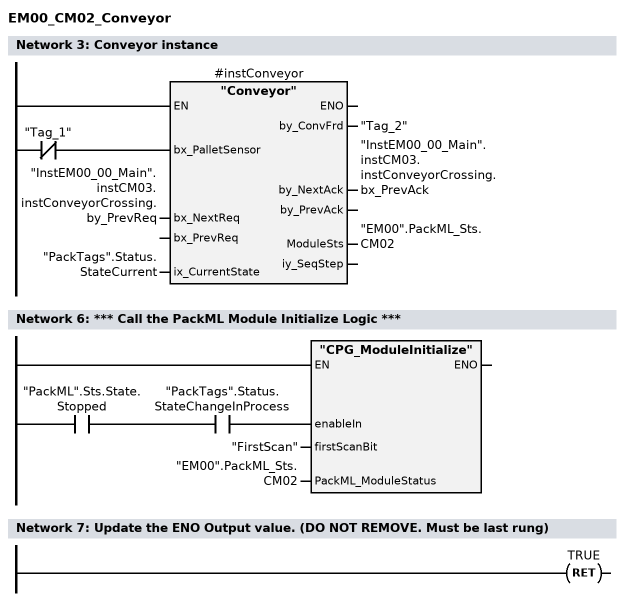
   RUNG wire#powerrail
      #instConveyor(bx_PalletSensor := wire#w1, bx_NextReq := "InstEM00_00_Main".instCM03.instConveyorCrossing.by_PrevReq, bx_PrevReq :=, ix_CurrentState := "PackTags".Status.StateCurrent, by_ConvFrd => "Tag_2", by_NextAck => "InstEM00_00_Main".instCM03.instConveyorCrossing.bx_PrevAck, by_PrevAck =>, ModuleSts => "EM00".PackML_Sts.CM02, iy_SeqStep =>)
   END_RUNG
   RUNG wire#powerrail
      I_Contact( "Tag_1" )
   END_RUNG wire#w1
   // the same network as SCL:
   #instConveyor(bx_PalletSensor := NOT "Tag_1",   // "Conveyor"
                 bx_NextReq := "InstEM00_00_Main".instCM03.instConveyorCrossing.by_PrevReq,
                 ix_CurrentState := "PackTags".Status.StateCurrent,
                 by_ConvFrd => "Tag_2",
                 by_NextAck => "InstEM00_00_Main".instCM03.instConveyorCrossing.bx_PrevAck,
                 ModuleSts => "EM00".PackML_Sts.CM02);
END_REGION

REGION Network 4: *** Begin the Event Information Section ***
END_REGION

REGION Network 5: *** Begin the State Model Status Feedback Section ***
END_REGION

REGION Network 6: *** Call the PackML Module Initialize Logic ***
   RUNG wire#powerrail
      "CPG_ModuleInitialize"(enableIn := wire#w1, firstScanBit := "FirstScan", PackML_ModuleStatus := "EM00".PackML_Sts.CM02)
   END_RUNG
   RUNG wire#powerrail
      Contact( "PackML".Sts.State.Stopped )
      Contact( "PackTags".Status.StateChangeInProcess )
   END_RUNG wire#w1
   // the same network as SCL:
   "CPG_ModuleInitialize"(enableIn := "PackML".Sts.State.Stopped AND "PackTags".Status.StateChangeInProcess,
                          firstScanBit := "FirstScan",
                          PackML_ModuleStatus := "EM00".PackML_Sts.CM02);
END_REGION

REGION Network 7: Update the ENO Output value. (DO NOT REMOVE. Must be last rung)
   RUNG wire#powerrail
      ReturnCoil( TRUE )
   END_RUNG
   // the same network as SCL:
   ENO := TRUE;
   RETURN;
END_REGION
END_FUNCTION_BLOCK

FUNCTION_BLOCK "EM00_CM03_ConveyorCrossing"   // FB31653, LAD
TITLE = EM00_CM03
{ S7_Optimized_Access := 'TRUE' }
AUTHOR : tech.team.motioncontrol@siemens.com
FAMILY : CPG
VERSION : 1.1
// Support: tech.team.motioncontrol@siemens.com
   VAR
      statDummyBool : Bool;   // dummy bool - placeholder
      instConveyorCrossing : "ConveyorCrossing";
   END_VAR
BEGIN

REGION Network 1: *** Begin the Setpoint Management Information Section ***
END_REGION

REGION Network 2: *** Begin the Logic Section ***
END_REGION

REGION Network 3: Conveyor crossing instance
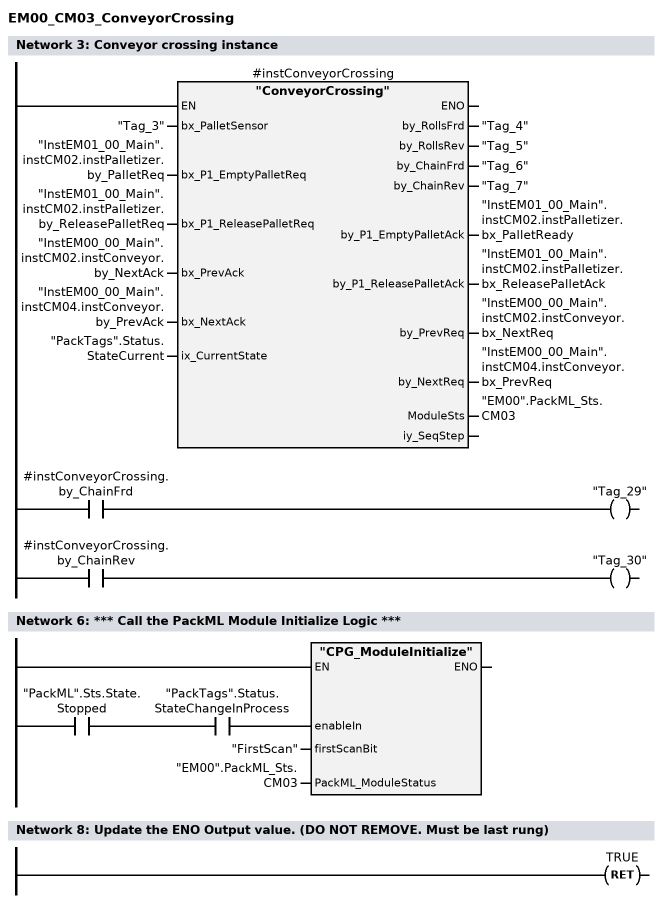
   RUNG wire#powerrail
      #instConveyorCrossing(bx_PalletSensor := "Tag_3", bx_P1_EmptyPalletReq := "InstEM01_00_Main".instCM02.instPalletizer.by_PalletReq, bx_P1_ReleasePalletReq := "InstEM01_00_Main".instCM02.instPalletizer.by_ReleasePalletReq, bx_PrevAck := "InstEM00_00_Main".instCM02.instConveyor.by_NextAck, bx_NextAck := "InstEM00_00_Main".instCM04.instConveyor.by_PrevAck, ix_CurrentState := "PackTags".Status.StateCurrent, by_RollsFrd => "Tag_4", by_RollsRev => "Tag_5", by_ChainFrd => "Tag_6", by_ChainRev => "Tag_7", by_P1_EmptyPalletAck => "InstEM01_00_Main".instCM02.instPalletizer.bx_PalletReady, by_P1_ReleasePalletAck => "InstEM01_00_Main".instCM02.instPalletizer.bx_ReleasePalletAck, by_PrevReq => "InstEM00_00_Main".instCM02.instConveyor.bx_NextReq, by_NextReq => "InstEM00_00_Main".instCM04.instConveyor.bx_PrevReq, ModuleSts => "EM00".PackML_Sts.CM03, iy_SeqStep =>)
   END_RUNG
   RUNG wire#powerrail
      Contact( #instConveyorCrossing.by_ChainFrd )
      Coil( "Tag_29" )
   END_RUNG
   RUNG wire#powerrail
      Contact( #instConveyorCrossing.by_ChainRev )
      Coil( "Tag_30" )
   END_RUNG
   // the same network as SCL:
   #instConveyorCrossing(bx_PalletSensor := "Tag_3",   // "ConveyorCrossing"
                         bx_P1_EmptyPalletReq := "InstEM01_00_Main".instCM02.instPalletizer.by_PalletReq,
                         bx_P1_ReleasePalletReq := "InstEM01_00_Main".instCM02.instPalletizer.by_ReleasePalletReq,
                         bx_PrevAck := "InstEM00_00_Main".instCM02.instConveyor.by_NextAck,
                         bx_NextAck := "InstEM00_00_Main".instCM04.instConveyor.by_PrevAck,
                         ix_CurrentState := "PackTags".Status.StateCurrent,
                         by_RollsFrd => "Tag_4",
                         by_RollsRev => "Tag_5",
                         by_ChainFrd => "Tag_6",
                         by_ChainRev => "Tag_7",
                         by_P1_EmptyPalletAck => "InstEM01_00_Main".instCM02.instPalletizer.bx_PalletReady,
                         by_P1_ReleasePalletAck => "InstEM01_00_Main".instCM02.instPalletizer.bx_ReleasePalletAck,
                         by_PrevReq => "InstEM00_00_Main".instCM02.instConveyor.bx_NextReq,
                         by_NextReq => "InstEM00_00_Main".instCM04.instConveyor.bx_PrevReq,
                         ModuleSts => "EM00".PackML_Sts.CM03);
   "Tag_29" := #instConveyorCrossing.by_ChainFrd;
   "Tag_30" := #instConveyorCrossing.by_ChainRev;
END_REGION

REGION Network 4: *** Begin the Event Information Section ***
END_REGION

REGION Network 5: *** Begin the State Model Status Feedback Section ***
END_REGION

REGION Network 6: *** Call the PackML Module Initialize Logic ***
   RUNG wire#powerrail
      "CPG_ModuleInitialize"(enableIn := wire#w1, firstScanBit := "FirstScan", PackML_ModuleStatus := "EM00".PackML_Sts.CM03)
   END_RUNG
   RUNG wire#powerrail
      Contact( "PackML".Sts.State.Stopped )
      Contact( "PackTags".Status.StateChangeInProcess )
   END_RUNG wire#w1
   // the same network as SCL:
   "CPG_ModuleInitialize"(enableIn := "PackML".Sts.State.Stopped AND "PackTags".Status.StateChangeInProcess,
                          firstScanBit := "FirstScan",
                          PackML_ModuleStatus := "EM00".PackML_Sts.CM03);
END_REGION

REGION Network 8: Update the ENO Output value. (DO NOT REMOVE. Must be last rung)
   RUNG wire#powerrail
      ReturnCoil( TRUE )
   END_RUNG
   // the same network as SCL:
   ENO := TRUE;
   RETURN;
END_REGION
END_FUNCTION_BLOCK

FUNCTION_BLOCK "EM00_CM04_Conveyor"   // FB31654, LAD
TITLE = EM00_CM04
{ S7_Optimized_Access := 'TRUE' }
AUTHOR : tech.team.motioncontrol@siemens.com
FAMILY : CPG
VERSION : 1.1
// Support: tech.team.motioncontrol@siemens.com
   VAR
      statDummyBool : Bool;   // dummy bool - placeholder
      instConveyor : "Conveyor";
   END_VAR
BEGIN

REGION Network 1: *** Begin the Setpoint Management Information Section ***
END_REGION

REGION Network 2: *** Begin the Logic Section ***
END_REGION

REGION Network 3: Conveyor instance
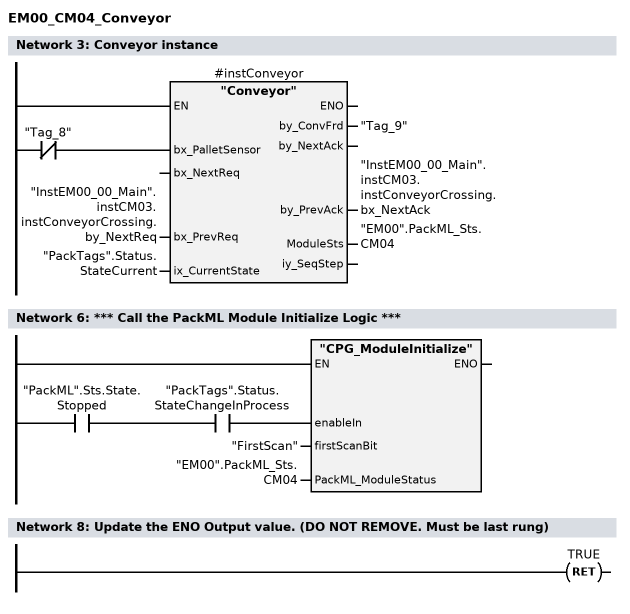
   RUNG wire#powerrail
      #instConveyor(bx_PalletSensor := wire#w1, bx_NextReq :=, bx_PrevReq := "InstEM00_00_Main".instCM03.instConveyorCrossing.by_NextReq, ix_CurrentState := "PackTags".Status.StateCurrent, by_ConvFrd => "Tag_9", by_NextAck =>, by_PrevAck => "InstEM00_00_Main".instCM03.instConveyorCrossing.bx_NextAck, ModuleSts => "EM00".PackML_Sts.CM04, iy_SeqStep =>)
   END_RUNG
   RUNG wire#powerrail
      I_Contact( "Tag_8" )
   END_RUNG wire#w1
   // the same network as SCL:
   #instConveyor(bx_PalletSensor := NOT "Tag_8",   // "Conveyor"
                 bx_PrevReq := "InstEM00_00_Main".instCM03.instConveyorCrossing.by_NextReq,
                 ix_CurrentState := "PackTags".Status.StateCurrent,
                 by_ConvFrd => "Tag_9",
                 by_PrevAck => "InstEM00_00_Main".instCM03.instConveyorCrossing.bx_NextAck,
                 ModuleSts => "EM00".PackML_Sts.CM04);
END_REGION

REGION Network 4: *** Begin the Event Information Section ***
END_REGION

REGION Network 5: *** Begin the State Model Status Feedback Section ***
END_REGION

REGION Network 6: *** Call the PackML Module Initialize Logic ***
   RUNG wire#powerrail
      "CPG_ModuleInitialize"(enableIn := wire#w1, firstScanBit := "FirstScan", PackML_ModuleStatus := "EM00".PackML_Sts.CM04)
   END_RUNG
   RUNG wire#powerrail
      Contact( "PackML".Sts.State.Stopped )
      Contact( "PackTags".Status.StateChangeInProcess )
   END_RUNG wire#w1
   // the same network as SCL:
   "CPG_ModuleInitialize"(enableIn := "PackML".Sts.State.Stopped AND "PackTags".Status.StateChangeInProcess,
                          firstScanBit := "FirstScan",
                          PackML_ModuleStatus := "EM00".PackML_Sts.CM04);
END_REGION

REGION Network 8: Update the ENO Output value. (DO NOT REMOVE. Must be last rung)
   RUNG wire#powerrail
      ReturnCoil( TRUE )
   END_RUNG
   // the same network as SCL:
   ENO := TRUE;
   RETURN;
END_REGION
END_FUNCTION_BLOCK

FUNCTION_BLOCK "EM00_CM05_ConveyorCrossing"   // FB31655, LAD
TITLE = EM00_CM05
{ S7_Optimized_Access := 'TRUE' }
AUTHOR : tech.team.motioncontrol@siemens.com
FAMILY : CPG
VERSION : 1.1
// Support: tech.team.motioncontrol@siemens.com
   VAR
      statDummyBool : Bool;   // dummy bool - placeholder
   END_VAR
BEGIN

REGION Network 1: *** Begin the Setpoint Management Information Section ***
END_REGION

REGION Network 2: *** Begin the Logic Section ***
END_REGION

REGION Network 3: *** Begin the Event Information Section ***
END_REGION

REGION Network 4: *** Begin the State Model Status Feedback Section ***
END_REGION

REGION Network 5: *** Call the PackML Module Initialize Logic ***
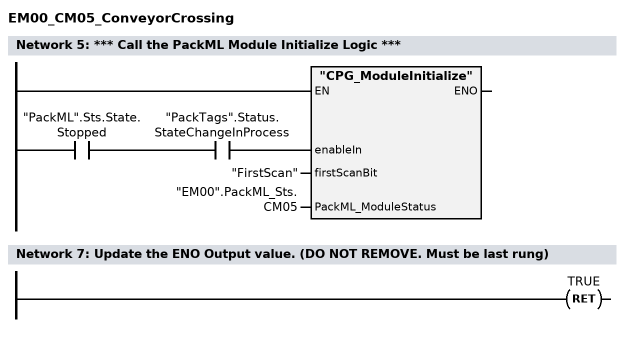
   RUNG wire#powerrail
      "CPG_ModuleInitialize"(enableIn := wire#w1, firstScanBit := "FirstScan", PackML_ModuleStatus := "EM00".PackML_Sts.CM05)
   END_RUNG
   RUNG wire#powerrail
      Contact( "PackML".Sts.State.Stopped )
      Contact( "PackTags".Status.StateChangeInProcess )
   END_RUNG wire#w1
   // the same network as SCL:
   "CPG_ModuleInitialize"(enableIn := "PackML".Sts.State.Stopped AND "PackTags".Status.StateChangeInProcess,
                          firstScanBit := "FirstScan",
                          PackML_ModuleStatus := "EM00".PackML_Sts.CM05);
END_REGION

REGION Network 7: Update the ENO Output value. (DO NOT REMOVE. Must be last rung)
   RUNG wire#powerrail
      ReturnCoil( TRUE )
   END_RUNG
   // the same network as SCL:
   ENO := TRUE;
   RETURN;
END_REGION
END_FUNCTION_BLOCK

// folder: EM01_Palletizing

FUNCTION_BLOCK "EM01_00_Main"   // FB31660, LAD
TITLE = EM01_00_Main
{ S7_Optimized_Access := 'TRUE' }
AUTHOR : tech.team.motioncontrol@siemens.com
FAMILY : CPG
VERSION : 1.1
// Support: tech.team.motioncontrol@siemens.com
   VAR
      instEventControl : "EM01_01_EventControl";   // Instance DB - EM's Event Control Logic
      instPackML_ModuleSum : "EM01_02_PackML_ModuleSum";   // Instance DB - EM's PackML Module Summation Logic
      instCM01 : "EM01_CM01_Conveyor";   // Instance DB - CM01
      instCM02 : "EM01_CM02_Palletizer";   // Instance DB - CM02
   END_VAR
   VAR_TEMP   // added for the SCL form of the ladder/FBD networks
      _w1 : Bool;
   END_VAR
BEGIN

REGION Network 1: *** BEGIN MAIN LOGIC SECTION ***
END_REGION

REGION Network 2: Call the Control Module Logic - CM01
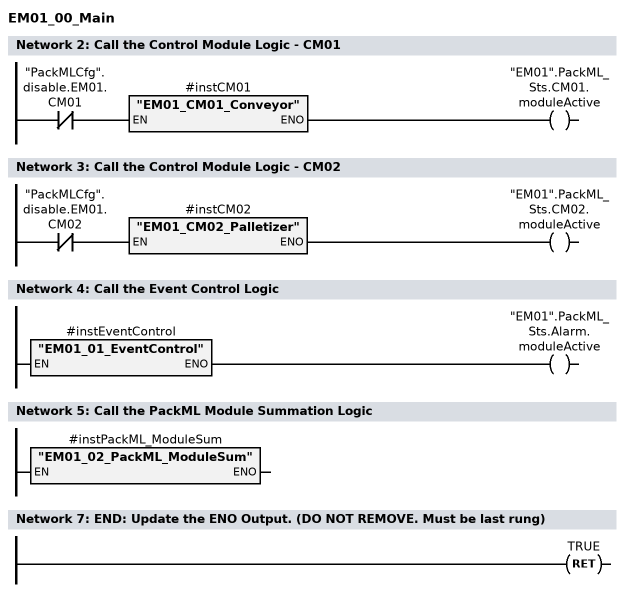
   RUNG wire#powerrail
      I_Contact( "PackMLCfg".disable.EM01.CM01 )
      #instCM01()
      Coil( "EM01".PackML_Sts.CM01.moduleActive )
   END_RUNG
   // the same network as SCL:
   #instCM01(EN := NOT "PackMLCfg".disable.EM01.CM01, ENO => #_w1);   // "EM01_CM01_Conveyor"
   "EM01".PackML_Sts.CM01.moduleActive := #_w1;
END_REGION

REGION Network 3: Call the Control Module Logic - CM02
   RUNG wire#powerrail
      I_Contact( "PackMLCfg".disable.EM01.CM02 )
      #instCM02()
      Coil( "EM01".PackML_Sts.CM02.moduleActive )
   END_RUNG
   // the same network as SCL:
   #instCM02(EN := NOT "PackMLCfg".disable.EM01.CM02, ENO => #_w1);   // "EM01_CM02_Palletizer"
   "EM01".PackML_Sts.CM02.moduleActive := #_w1;
END_REGION

REGION Network 4: Call the Event Control Logic
   RUNG wire#powerrail
      #instEventControl()
      Coil( "EM01".PackML_Sts.Alarm.moduleActive )
   END_RUNG
   // the same network as SCL:
   #instEventControl(ENO => #_w1);   // "EM01_01_EventControl"
   "EM01".PackML_Sts.Alarm.moduleActive := #_w1;
END_REGION

REGION Network 5: Call the PackML Module Summation Logic
   RUNG wire#powerrail
      #instPackML_ModuleSum()
   END_RUNG
   // the same network as SCL:
   #instPackML_ModuleSum();   // "EM01_02_PackML_ModuleSum"
END_REGION

REGION Network 7: END: Update the ENO Output. (DO NOT REMOVE. Must be last rung)
   RUNG wire#powerrail
      ReturnCoil( TRUE )
   END_RUNG
   // the same network as SCL:
   ENO := TRUE;
   RETURN;
END_REGION
END_FUNCTION_BLOCK

FUNCTION_BLOCK "EM01_01_EventControl"   // FB31661, LAD
TITLE = EM01_01_EventControl
{ S7_Optimized_Access := 'TRUE' }
AUTHOR : tech.team.motioncontrol@siemens.com
FAMILY : CPG
VERSION : 1.1
// Support: tech.team.motioncontrol@siemens.com
   VAR
      instEventMgr_Alarm : "CPG_EventManager";   // instance FB - Event Manager - Alarm Events
      instEventMgr_Warning : "CPG_EventManager";   // instance FB - Event Manager - Warning Events
      instEventMgr_Status : "CPG_EventManager";   // instance FB - Event Manager - Status Events
      instStatus_AlarmNotReset : "CPG_Event";   // instance FB - PackML Event - Alarms not reset
      statEventMgr_Cmd_Reset : Bool;   // Reset Cmd for all event managers
      statEventMgr_Cmd_Clear1stFlt : Bool;   // Clear 1st Fault Cmd for all event managers
      statEventMgr_Clear1stFlt_OS : Bool;   // Clear 1st Fault Cmd - One shot
   END_VAR
   VAR_TEMP   // added for the SCL form of the ladder/FBD networks
      _w1 : Bool;
      _w2 : Bool;
   END_VAR
BEGIN

REGION Network 1: ** STATE MODEL REPORTING STATUS ****
END_REGION

REGION Network 2: *** Call the PackML Module Initialize Logic ***
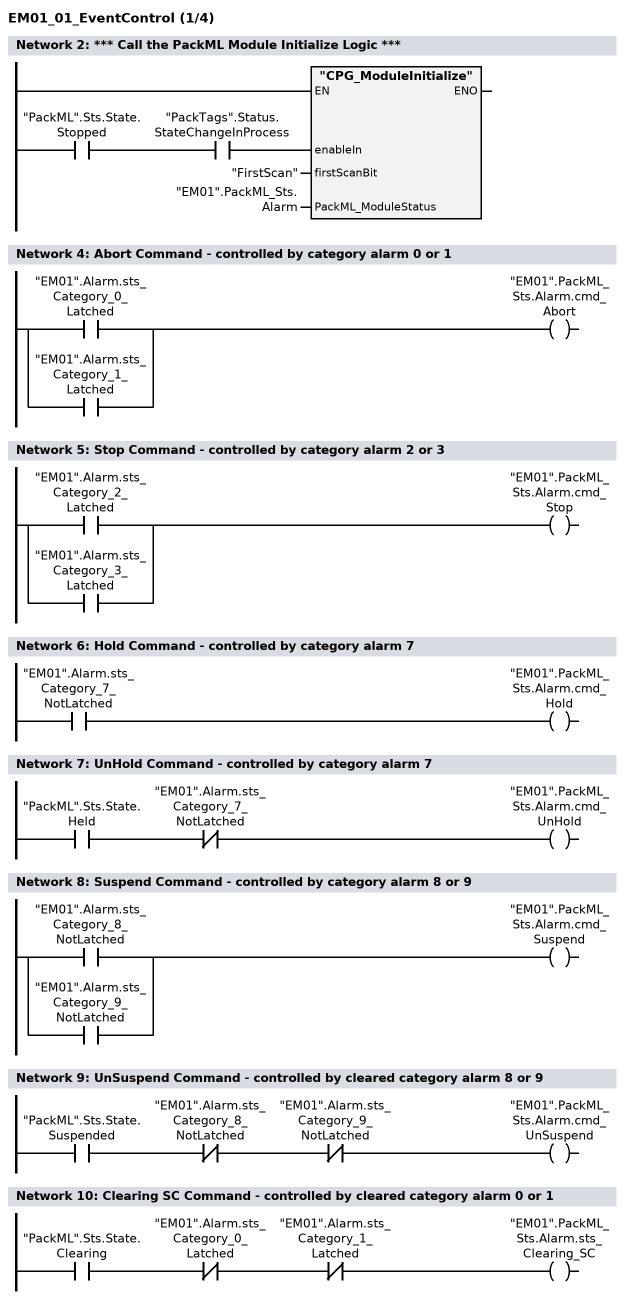
   RUNG wire#powerrail
      "CPG_ModuleInitialize"(enableIn := wire#w1, firstScanBit := "FirstScan", PackML_ModuleStatus := "EM01".PackML_Sts.Alarm)
   END_RUNG
   RUNG wire#powerrail
      Contact( "PackML".Sts.State.Stopped )
      Contact( "PackTags".Status.StateChangeInProcess )
   END_RUNG wire#w1
   // the same network as SCL:
   "CPG_ModuleInitialize"(enableIn := "PackML".Sts.State.Stopped AND "PackTags".Status.StateChangeInProcess,
                          firstScanBit := "FirstScan",
                          PackML_ModuleStatus := "EM01".PackML_Sts.Alarm);
END_REGION

REGION Network 3: Begin the LOGIC section.
END_REGION

REGION Network 4: Abort Command - controlled by category alarm 0 or 1
   RUNG wire#powerrail
      Contact( "EM01".Alarm.sts_Category_0_Latched )
      wire#w1
      Coil( "EM01".PackML_Sts.Alarm.cmd_Abort )
   END_RUNG
   RUNG wire#powerrail
      Contact( "EM01".Alarm.sts_Category_1_Latched )
   END_RUNG wire#w1
   // the same network as SCL:
   "EM01".PackML_Sts.Alarm.cmd_Abort := "EM01".Alarm.sts_Category_0_Latched OR "EM01".Alarm.sts_Category_1_Latched;
END_REGION

REGION Network 5: Stop Command - controlled by category alarm 2 or 3
   RUNG wire#powerrail
      Contact( "EM01".Alarm.sts_Category_2_Latched )
      wire#w1
      Coil( "EM01".PackML_Sts.Alarm.cmd_Stop )
   END_RUNG
   RUNG wire#powerrail
      Contact( "EM01".Alarm.sts_Category_3_Latched )
   END_RUNG wire#w1
   // the same network as SCL:
   "EM01".PackML_Sts.Alarm.cmd_Stop := "EM01".Alarm.sts_Category_2_Latched OR "EM01".Alarm.sts_Category_3_Latched;
END_REGION

REGION Network 6: Hold Command - controlled by category alarm 7
   RUNG wire#powerrail
      Contact( "EM01".Alarm.sts_Category_7_NotLatched )
      Coil( "EM01".PackML_Sts.Alarm.cmd_Hold )
   END_RUNG
   // the same network as SCL:
   "EM01".PackML_Sts.Alarm.cmd_Hold := "EM01".Alarm.sts_Category_7_NotLatched;
END_REGION

REGION Network 7: UnHold Command - controlled by category alarm 7
   RUNG wire#powerrail
      Contact( "PackML".Sts.State.Held )
      I_Contact( "EM01".Alarm.sts_Category_7_NotLatched )
      Coil( "EM01".PackML_Sts.Alarm.cmd_UnHold )
   END_RUNG
   // the same network as SCL:
   "EM01".PackML_Sts.Alarm.cmd_UnHold := "PackML".Sts.State.Held AND NOT "EM01".Alarm.sts_Category_7_NotLatched;
END_REGION

REGION Network 8: Suspend Command - controlled by category alarm 8 or 9
   RUNG wire#powerrail
      Contact( "EM01".Alarm.sts_Category_8_NotLatched )
      wire#w1
      Coil( "EM01".PackML_Sts.Alarm.cmd_Suspend )
   END_RUNG
   RUNG wire#powerrail
      Contact( "EM01".Alarm.sts_Category_9_NotLatched )
   END_RUNG wire#w1
   // the same network as SCL:
   "EM01".PackML_Sts.Alarm.cmd_Suspend := "EM01".Alarm.sts_Category_8_NotLatched OR "EM01".Alarm.sts_Category_9_NotLatched;
END_REGION

REGION Network 9: UnSuspend Command - controlled by cleared category alarm 8 or 9
   RUNG wire#powerrail
      Contact( "PackML".Sts.State.Suspended )
      I_Contact( "EM01".Alarm.sts_Category_8_NotLatched )
      I_Contact( "EM01".Alarm.sts_Category_9_NotLatched )
      Coil( "EM01".PackML_Sts.Alarm.cmd_UnSuspend )
   END_RUNG
   // the same network as SCL:
   "EM01".PackML_Sts.Alarm.cmd_UnSuspend := "PackML".Sts.State.Suspended AND NOT "EM01".Alarm.sts_Category_8_NotLatched AND NOT "EM01".Alarm.sts_Category_9_NotLatched;
END_REGION

REGION Network 10: Clearing SC Command - controlled by cleared category alarm 0 or 1
   RUNG wire#powerrail
      Contact( "PackML".Sts.State.Clearing )
      I_Contact( "EM01".Alarm.sts_Category_0_Latched )
      I_Contact( "EM01".Alarm.sts_Category_1_Latched )
      Coil( "EM01".PackML_Sts.Alarm.sts_Clearing_SC )
   END_RUNG
   // the same network as SCL:
   "EM01".PackML_Sts.Alarm.sts_Clearing_SC := "PackML".Sts.State.Clearing AND NOT "EM01".Alarm.sts_Category_0_Latched AND NOT "EM01".Alarm.sts_Category_1_Latched;
END_REGION

REGION Network 11: Resetting SC Command - controlled by cleared category alarm 0-3
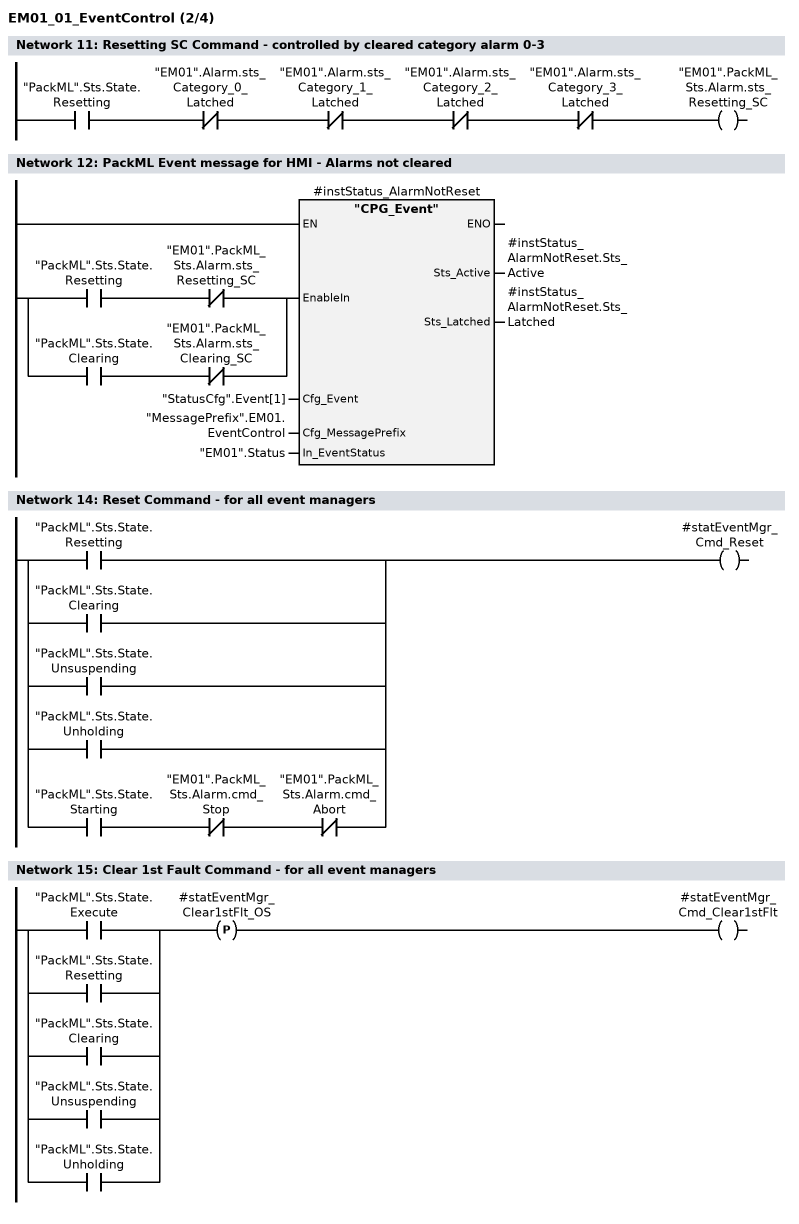
   RUNG wire#powerrail
      Contact( "PackML".Sts.State.Resetting )
      I_Contact( "EM01".Alarm.sts_Category_0_Latched )
      I_Contact( "EM01".Alarm.sts_Category_1_Latched )
      I_Contact( "EM01".Alarm.sts_Category_2_Latched )
      I_Contact( "EM01".Alarm.sts_Category_3_Latched )
      Coil( "EM01".PackML_Sts.Alarm.sts_Resetting_SC )
   END_RUNG
   // the same network as SCL:
   "EM01".PackML_Sts.Alarm.sts_Resetting_SC := "PackML".Sts.State.Resetting AND NOT "EM01".Alarm.sts_Category_0_Latched AND NOT "EM01".Alarm.sts_Category_1_Latched AND NOT "EM01".Alarm.sts_Category_2_Latched AND NOT "EM01".Alarm.sts_Category_3_Latched;
END_REGION

REGION Network 12: PackML Event message for HMI - Alarms not cleared
   RUNG wire#powerrail
      #instStatus_AlarmNotReset(EnableIn := wire#w1, Cfg_Event := "StatusCfg".Event[1], Cfg_MessagePrefix := "MessagePrefix".EM01.EventControl, In_EventStatus := "EM01".Status, Sts_Active => #instStatus_AlarmNotReset.Sts_Active, Sts_Latched => #instStatus_AlarmNotReset.Sts_Latched)
   END_RUNG
   RUNG wire#powerrail
      Contact( "PackML".Sts.State.Resetting )
      I_Contact( "EM01".PackML_Sts.Alarm.sts_Resetting_SC )
   END_RUNG wire#w1
   RUNG wire#powerrail
      Contact( "PackML".Sts.State.Clearing )
      I_Contact( "EM01".PackML_Sts.Alarm.sts_Clearing_SC )
   END_RUNG wire#w1
   // the same network as SCL:
   #instStatus_AlarmNotReset(EnableIn := ("PackML".Sts.State.Resetting AND NOT "EM01".PackML_Sts.Alarm.sts_Resetting_SC) OR ("PackML".Sts.State.Clearing AND NOT "EM01".PackML_Sts.Alarm.sts_Clearing_SC),   // "CPG_Event"
                           Cfg_Event := "StatusCfg".Event[1],
                           Cfg_MessagePrefix := "MessagePrefix".EM01.EventControl,
                           In_EventStatus := "EM01".Status,
                           Sts_Active => #instStatus_AlarmNotReset.Sts_Active,
                           Sts_Latched => #instStatus_AlarmNotReset.Sts_Latched);
END_REGION

REGION Network 13: *** EVENT CONTROL MANAGERS ***
END_REGION

REGION Network 14: Reset Command - for all event managers
   RUNG wire#powerrail
      Contact( "PackML".Sts.State.Resetting )
      wire#w1
      Coil( #statEventMgr_Cmd_Reset )
   END_RUNG
   RUNG wire#powerrail
      Contact( "PackML".Sts.State.Clearing )
   END_RUNG wire#w1
   RUNG wire#powerrail
      Contact( "PackML".Sts.State.Unsuspending )
   END_RUNG wire#w1
   RUNG wire#powerrail
      Contact( "PackML".Sts.State.Unholding )
   END_RUNG wire#w1
   RUNG wire#powerrail
      Contact( "PackML".Sts.State.Starting )
      I_Contact( "EM01".PackML_Sts.Alarm.cmd_Stop )
      I_Contact( "EM01".PackML_Sts.Alarm.cmd_Abort )
   END_RUNG wire#w1
   // the same network as SCL:
   #statEventMgr_Cmd_Reset := "PackML".Sts.State.Resetting OR "PackML".Sts.State.Clearing OR "PackML".Sts.State.Unsuspending OR "PackML".Sts.State.Unholding OR ("PackML".Sts.State.Starting AND NOT "EM01".PackML_Sts.Alarm.cmd_Stop AND NOT "EM01".PackML_Sts.Alarm.cmd_Abort);
END_REGION

REGION Network 15: Clear 1st Fault Command - for all event managers
   RUNG wire#powerrail
      Contact( "PackML".Sts.State.Execute )
      wire#w1
      P_Trig( #statEventMgr_Clear1stFlt_OS )
      Coil( #statEventMgr_Cmd_Clear1stFlt )
   END_RUNG
   RUNG wire#powerrail
      Contact( "PackML".Sts.State.Resetting )
   END_RUNG wire#w1
   RUNG wire#powerrail
      Contact( "PackML".Sts.State.Clearing )
   END_RUNG wire#w1
   RUNG wire#powerrail
      Contact( "PackML".Sts.State.Unsuspending )
   END_RUNG wire#w1
   RUNG wire#powerrail
      Contact( "PackML".Sts.State.Unholding )
   END_RUNG wire#w1
   // the same network as SCL:
   #_w1 := "PackML".Sts.State.Execute OR "PackML".Sts.State.Resetting OR "PackML".Sts.State.Clearing OR "PackML".Sts.State.Unsuspending OR "PackML".Sts.State.Unholding;
   #_w2 := #_w1 AND NOT #statEventMgr_Clear1stFlt_OS;   // rising edge
   #statEventMgr_Clear1stFlt_OS := #_w1;
   #statEventMgr_Cmd_Clear1stFlt := #_w2;
END_REGION

REGION Network 16: Call the Event Manager logic for EM alarms
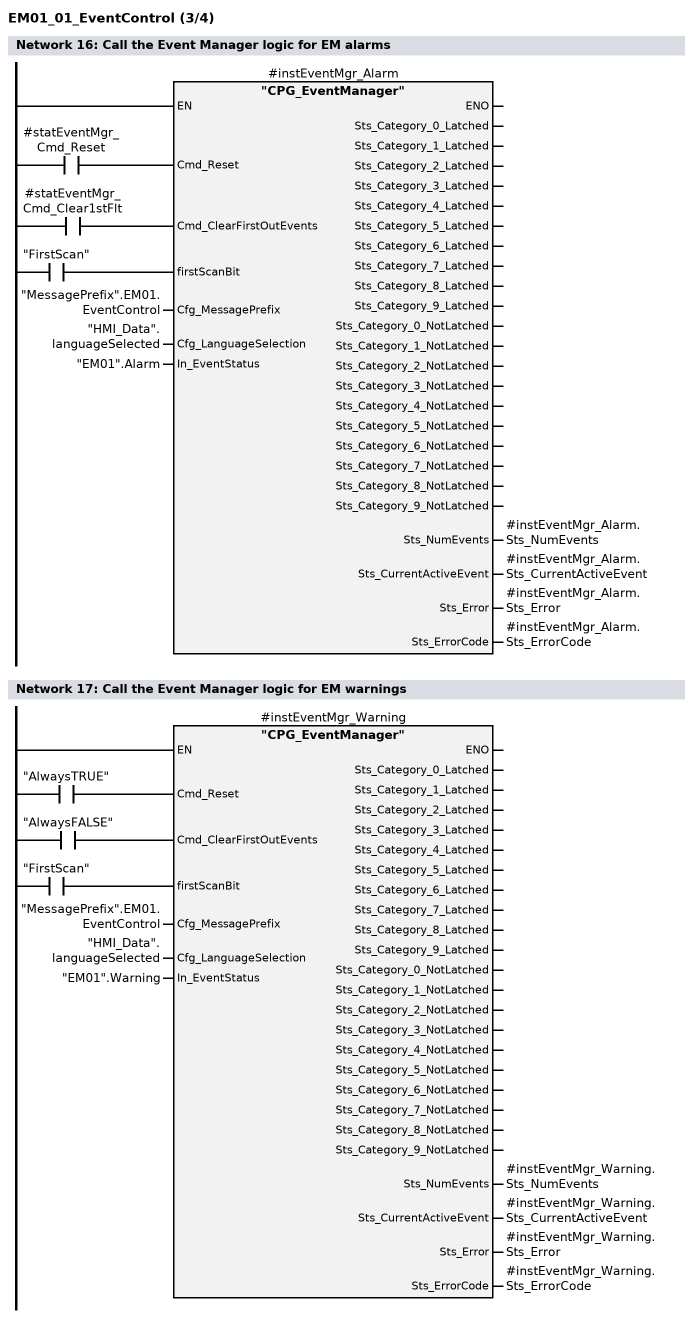
   RUNG wire#powerrail
      #instEventMgr_Alarm(Cmd_Reset := wire#w1, Cmd_ClearFirstOutEvents := wire#w2, firstScanBit := wire#w3, Cfg_MessagePrefix := "MessagePrefix".EM01.EventControl, Cfg_LanguageSelection := "HMI_Data".languageSelected, In_EventStatus := "EM01".Alarm, Sts_Category_0_Latched =>, Sts_Category_1_Latched =>, Sts_Category_2_Latched =>, Sts_Category_3_Latched =>, Sts_Category_4_Latched =>, Sts_Category_5_Latched =>, Sts_Category_6_Latched =>, Sts_Category_7_Latched =>, Sts_Category_8_Latched =>, Sts_Category_9_Latched =>, Sts_Category_0_NotLatched =>, Sts_Category_1_NotLatched =>, Sts_Category_2_NotLatched =>, Sts_Category_3_NotLatched =>, Sts_Category_4_NotLatched =>, Sts_Category_5_NotLatched =>, Sts_Category_6_NotLatched =>, Sts_Category_7_NotLatched =>, Sts_Category_8_NotLatched =>, Sts_Category_9_NotLatched =>, Sts_NumEvents => #instEventMgr_Alarm.Sts_NumEvents, Sts_CurrentActiveEvent => #instEventMgr_Alarm.Sts_CurrentActiveEvent, Sts_Error => #instEventMgr_Alarm.Sts_Error, Sts_ErrorCode => #instEventMgr_Alarm.Sts_ErrorCode)
   END_RUNG
   RUNG wire#powerrail
      Contact( #statEventMgr_Cmd_Reset )
   END_RUNG wire#w1
   RUNG wire#powerrail
      Contact( #statEventMgr_Cmd_Clear1stFlt )
   END_RUNG wire#w2
   RUNG wire#powerrail
      Contact( "FirstScan" )
   END_RUNG wire#w3
   // the same network as SCL:
   #instEventMgr_Alarm(Cmd_Reset := #statEventMgr_Cmd_Reset,   // "CPG_EventManager"
                       Cmd_ClearFirstOutEvents := #statEventMgr_Cmd_Clear1stFlt,
                       firstScanBit := "FirstScan",